// Mitsubishi GX Works2 project: 70常温静置库1130   PLC: Q10UDEH (continued)
IF NOT m_xInitial THEN
	ConveyorMotor.tLoadDelay:=T#100ms;
	ConveyorMotor.tUnloadAlarmDelay:=T#30s;
	ConveyorMotor.xPosLimit:=1;
	ConveyorMotor.xNegLimit:=1;
	ConveyorMotor.xSizeDeficientDetect:=0;
	ConveyorMotor.xZoneClear:=0;
	ConveyorMotor.tZoneClearTime:=T#10s;
	m_xInitial:=1;
END_IF;
(*//自动
//复位信号把步号置0，但xLoad与xUnload没有复位，调用程序需要注意复位后把这两个信号置零，以免发生误动作
//物料有无判断增加延时，防止开自动瞬间误动作发生*)
m_tonPresentDelay(IN:= ConveyorMotor.xCWPresent OR ConveyorMotor.xCCWPresent,
                  PT:=T#100ms,
				  Q:= m_xPresentDelay,
				  ET:= m_tPresentDelayCurrentTime);

CASE iStep OF
	0:(*//初始化*)
	ConveyorMotor.xMotorCW:=0;
	ConveyorMotor.xMotorCCW:=0;
	ConveyorMotor.iProductCategoryOut:=0;
(*	//判断物料有无传感器*)	
		IF m_xPresentDelay THEN			
			ConveyorMotor.xEmpty:=0;
			IF g_xAuto AND NOT ConveyorMotor.xError THEN(*//自动情况下进行跳转*)(*无超限报警*)
				iStep:=3;
			END_IF;
		ELSE
			ConveyorMotor.xEmpty:=1;
			IF g_xAuto AND NOT ConveyorMotor.xError THEN(*//自动情况下进行跳转*)(*无超限报警*)
				iStep:=1;	
			END_IF;		
	END_IF;	
	1: (*//上料*)
	ConveyorMotor.xNextRun:=0;
	IF ConveyorMotor.xLoad    THEN (*//上料开始*)
		ConveyorMotor.iProductCategory:=0;	(*//上料开始清除产品信息*)
		iStep:=2;		
	END_IF;
	2: (*//上料完成*)
	IF ConveyorMotor.iProductCategoryIn<>0 THEN
		ConveyorMotor.iProductCategory:=ConveyorMotor.iProductCategoryIn;(* //产品信息传入*)
	END_IF;
	IF ConveyorMotor.xloadCCW THEN
		ConveyorMotor.xMotorCCW:=1; 
		ConveyorMotor.xMotorCW:=0;
	ELSE
	    ConveyorMotor.xMotorCW:=1;  
		ConveyorMotor.xMotorCCW:=0;
	END_IF;
		m_tonLoadDelay(IN:= (ConveyorMotor.xCWPresent AND NOT ConveyorMotor.xloadCCW) 
		                                        OR (ConveyorMotor.xCCWPresent AND ConveyorMotor.xloadCCW) ,
		                               PT:= ConveyorMotor.tLoadDelay ,
		                               Q:= m_xLoadDelayOut ,
		                               ET:= m_tLoadTimer );
	    IF m_xLoadDelayOut THEN 	 
		    iStep:=3;
		END_IF;
	3:(*//下料请求*)	
	ConveyorMotor.xMotorCW:=0;
	ConveyorMotor.xMotorCCW:=0;
	ConveyorMotor.xEmpty:=0;
	IF ConveyorMotor.xUnload AND NOT ConveyorMotor.xOverWidthAlarm  THEN (*无超宽报警可以下料*)
		iStep:=4;
	END_IF;
	4:(*	//下料完成*)
	IF ConveyorMotor.xUnloadCCW THEN   
		ConveyorMotor.xMotorCCW:=1;  
		ConveyorMotor.xMotorCW:=0;
		ELSE
	    ConveyorMotor.xMotorCW:=1;  
		ConveyorMotor.xMotorCCW:=0;
	END_IF;
	ConveyorMotor.xNextRun:=1; (*下一段线体旋转*)
	ConveyorMotor.iProductCategoryOut:=ConveyorMotor.iProductCategory;(*产品型号输出给下一段线体*)
	IF NOT ConveyorMotor.xUnload THEN 
		istep:=0;
	END_IF;
END_CASE;
(*In-feed zone clear and ready to accept a load from upstream Conveyor*)
IF ldp(TRUE,g_xAuto) THEN
	m_xAutoClear:=1;
END_IF;
IF ldf(TRUE,g_xAuto) THEN
	m_xAutoClear:=0;
END_IF;
m_tonZoneClear(IN:= m_xAutoClear AND ConveyorMotor.xZoneClear ,PT:= ConveyorMotor.tZoneClearTime ,Q:=m_xZoneClearDone ,ET:= m_tZoneClearCurrentTime );
IF  m_xAutoClear AND ConveyorMotor.xZoneClear THEN
		ConveyorMotor.xMotorCW:=1; 
		iStep:=0;
END_IF;
IF ldf(TRUE, m_xAutoClear )THEN
	ConveyorMotor.xMotorCW:=0; 
END_IF;
IF NOT m_xAutoClear OR m_xZoneClearDone OR m_xPresentDelay THEN
	 m_xAutoClear:=0;
END_IF;	 
(*投入上料，搬出下料，也可用来初始化*)
IF LDP(TRUE,ConveyorMotor.xPutInto) THEN
	iStep:=0;
END_IF;
(*//当前任务显示*)
IF LDP(TRUE,ConveyorMotor.iDeviceID=g_iDeviceIDSelect) THEN
	g_iInsertTask:=ConveyorMotor.iProductCategory;
END_IF;
	(*//插入任务*)
IF g_xInsertTask AND ConveyorMotor.iDeviceID=g_iDeviceIDSelect THEN
	ConveyorMotor.iProductCategory:=g_iInsertTask;
END_IF;
(*//单线体复位，当设备号与本线体一致的时候执行复位*)
IF (g_xResetSingle AND ConveyorMotor.iDeviceID=g_iDeviceIDSelect)THEN (* //非正常情况下切断xNextRun不会复位，通过这个标志位会出发报警*)(*增加单体复位*)
	iStep:=0;
	ConveyorMotor.xNextRun:=0; 
	ConveyorMotor.xLimitAlarrm:=0;
	ConveyorMotor.xOverWidthAlarm:=0;
END_IF;
(*//手动*)
IF g_xManual THEN
(*	iStep:=0; *)(*//手动后上下料程序步骤清零*)
	(*//正转*)
	IF ConveyorMotor.xForward 
		AND ConveyorMotor.xBackward=0 
		AND ConveyorMotor.xMotorCCW=0 
		AND g_xEStop THEN
		ConveyorMotor.xMotorCW:=1;
		ConveyorMotor.xMotorCCW:=0;
		ELSE
		ConveyorMotor.xMotorCW:=0;
	END_IF;
	(*//反转*)
	IF ConveyorMotor.xBackward 
		AND ConveyorMotor.xForward=0 
		AND ConveyorMotor.xMotorCW=0 
		AND g_xEStop THEN
		ConveyorMotor.xMotorCCW:=1;
		conveyormotor.xMotorCW:=0;
		ELSE
		ConveyorMotor.xMotorCCW:=0;
	END_IF;
END_IF;
(*暂停*)
IF g_xPause THEN
	ConveyorMotor.xMotorCCW:=0;
	ConveyorMotor.xMotorCW:=0;
END_IF;
(*工作中信号输出*)
ConveyorMotor.xBusy:=ConveyorMotor.xMotorCCW OR ConveyorMotor.xMotorCW;
(*//未到达报警*)
m_tonNotArriveAlarm(IN:= iStep=0 AND ConveyorMotor.xNextRun  ,PT:= T#2s,Q:= ConveyorMotor.xNotArriveAlarm ,ET:= m_tNotArriveCurrentTime );
(*//下料超时报警*)
m_tonUnloadAlam(IN:= iStep=4,PT:=ConveyorMotor.tUnloadAlarmDelay,Q:= ConveyorMotor.xUnloadAlarm,ET:=m_tUnloadTimer );
(*//限位报警,进料检测开关失效*)
IF ( ((ConveyorMotor.xloadCCW AND NOT ConveyorMotor.xNegLimit)            (*反转上料，碰到负限位*)
	OR  ( NOT ConveyorMotor.xloadCCW AND NOT ConveyorMotor.xPosLimit)) (*正转上料，碰到正限位*)
    AND iStep=2) (*上料过程*)
    OR
   ( iStep=4 (*下料过程*)
	AND( (ConveyorMotor.xUnloadCCW AND NOT ConveyorMotor.xPosLimit)  
	OR (NOT ConveyorMotor.xUnloadCCW AND NOT ConveyorMotor.xNegLimit)))    
    THEN
    ConveyorMotor.xLimitAlarrm:=1;
    iStep:=0;
END_IF;
(*//超宽报警*)
IF (iStep=3 OR iStep=1) AND (NOT ConveyorMotor.xNegLimit OR NOT ConveyorMotor.xPosLimit) THEN
	ConveyorMotor.xOverWidthAlarm:=1;
END_IF;
(*//尺寸不足报警*)
(*//有料状态下检测两个开关都要有信号*)
IF iStep=3 AND ConveyorMotor.xSizeDeficientDetect AND (NOT ConveyorMotor.xCCWPresent OR NOT ConveyorMotor.xCWPresent)  THEN
	   ConveyorMotor.xOverWidthAlarm:=1;
	    iStep:=0;               
END_IF;
(*//总报警*)
ConveyorMotor.xError:=ConveyorMotor.xLimitAlarrm
                                              OR ConveyorMotor.xNotArriveAlarm
                                              OR ConveyorMotor.xUnloadAlarm                                             
                                              OR ConveyorMotor.xOverWidthAlarm;

(*//状态输出*)(*状态显示，容易造成指针容量不足*)
IF ConveyorMotor.xEmpty AND NOT ConveyorMotor.xBusy THEN
	m_wStateWord:=0;
END_IF;
IF ConveyorMotor.xEmpty=0 THEN
		m_wStateWord:=1;
END_IF;
IF ConveyorMotor.xBusy THEN
		m_wStateWord:=2;
END_IF;
IF ConveyorMotor.xLimitAlarrm THEN
		m_wStateWord:=3;
END_IF;
IF ConveyorMotor.xOverWidthAlarm THEN
		m_wStateWord:=4;
END_IF;
IF ConveyorMotor.xNotArriveAlarm THEN	
		m_wStateWord:=5;
END_IF;
IF ConveyorMotor.xUnloadAlarm THEN
		m_wStateWord:=6;	
END_IF;
(*选择本线体后，将状态赋值给全局变量进行显示*)
IF ConveyorMotor.iDeviceID=g_iDeviceIDSelect THEN
	g_iConveyorStatus:=m_wStateWord;
END_IF;
END_FUNCTION_BLOCK

FUNCTION_BLOCK DivideFolder
VAR_IN_OUT
  FolderIO : FolderIO;
  FolderConveyorIO : ConveyorIO;
END_VAR
VAR
  iFolderCount : INT;
  m_xInitial : BOOL;
  istep : INT;
  m_TONLoadDelay : TON;  (* 上料完成延时 *)
  m_xLoadDelay : BOOL;  (* 上料完成延时 *)
  m_tLoadDelay : TIME;  (* 上料完成延时 *)
  m_TONUpCylinderError : TON;
  m_tUpCylinderError : TIME;
  m_TONDownCylinderError : TON;
  m_tDownCylinderError : TIME;
  m_TONGrabCylinderError : TON;
  m_tGrabCylinderError : TIME;
END_VAR
VAR_INPUT
  i_xAuto : BOOL;  (* 自动 *)
END_VAR
(*拆盘机*)
(*Mr.Li修改2018.11.19调试*)
(*初始化*)
IF NOT m_xInitial  THEN
	FolderIO.i_iFloor:=3;
	 iFolderCount:=3;
	 	FolderIO.i_tSetOvertime:=T#5S;
		m_xInitial:=1;
END_IF;
(*自动*)
IF i_xAuto THEN
	FolderIO.o_xEntryPermit:=iFolderCount=3 AND FolderConveyorIO.xEmpty;(*线体状态为空且拆盘初始数量为3，才准上料*)
	m_TONLoadDelay(IN:= NOT FolderConveyorIO.xEmpty,
											PT:= T#100MS,
											Q:=m_xLoadDelay,
											ET:=m_tLoadDelay);

	CASE istep OF
		0:(*各种初始化*)
			FolderConveyorIO.xLoad:=0;
			FolderConveyorIO.xUnload:=0;
			FolderConveyorIO.xPutInto:=0;
			IF FolderConveyorIO.xEmpty THEN(*空的情况，0时上料，其他走流程*)
				IF iFolderCount=FolderIO.i_iFloor   THEN
					istep:=1; 					
				ELSE
					istep:=5;
				END_IF;	
			END_IF;		
			IF m_xLoadDelay THEN
				 IF FolderIO.i_xCylinderDownRetractDetect AND FolderIO.i_xCylinderUpRetractDetect THEN
					istep:=2;(*如果在1层，则顶起，需人为判断是否在指定位置，否则有翻框的危险*)
				ELSE
				 	istep:=3;(*如果有料不在1层，则抓紧，然后跳到第4步判断是否是叠盘，不是就放行*)
				 END_IF;
			END_IF;
		1:(*上料*)
			IF FolderIO.o_xEntryPermit THEN
				FolderConveyorIO.xLoad:=FolderIO.i_FrontConveyorNextRun;
			ELSE
				FolderConveyorIO.xLoad:=0;
			END_IF;(*有料等延时*)	
			IF m_xLoadDelay THEN
				iFolderCount:=FolderIO.i_iFloor;
				istep:=2;(**拆盘机顶起步骤*)
			END_IF;	
		2:(*上升至2层位置*)
				FolderIO.o_xCylinderDownRetract:=0;
				FolderIO.o_xCylinderDownExtend:=1;
				FolderIO.o_xCylinderUpRetract:=0;
				IF FolderIO.i_xCylinderDownExtendDetect   THEN
				istep:=3;
				END_IF;
		3:	(*夹紧夹爪*)
			IF FolderIO.i_xCylinderDownExtendDetect THEN
				FolderIO.o_xCylinderGrabExtend:=1;
				FolderIO.o_xCylinderGrabRetract:=0;
			END_IF;
			IF FolderIO.i_xCylinderGrabExtendDetect THEN
				istep:=4;
			END_IF;	
		4:(*再下降到1层，然后放行，在该位置判断是不是最后一次*)
				FolderIO.o_xCylinderUpRetract:=1;
				FolderIO.o_xCylinderUpExtend:=0;
				FolderIO.o_xCylinderDownRetract:=1;
				FolderIO.o_xCylinderDownExtend:=0;
				IF FolderIO.i_xCylinderDownRetractDetect AND FolderIO.i_xCylinderUpRetractDetect AND FolderIO.o_xExitPremit THEN
				FolderConveyorIO.xPutInto:=1;
				FolderConveyorIO.xUnload:=FolderIO.o_xExitPremit;
				ELSIF NOT FolderIO.i_xTrayDetect AND NOT FolderConveyorIO.xEmpty AND FolderIO.o_xExitPremit THEN 
						FolderConveyorIO.xUnload:=FolderIO.o_xExitPremit;
				ELSE 
					FolderConveyorIO.xPutInto:=0;
				FolderConveyorIO.xUnload:=0;
				END_IF;
					IF FolderIO.i_xCylinderDownRetractDetect AND FolderIO.i_xCylinderUpRetractDetect AND
						  FolderIO.i_xTrayDetect  AND  iFolderCount>0  AND ldp(TRUE,NOT  FolderConveyorIO.xUnload) THEN
						iFolderCount:=FolderIO.i_iFloor-1;					
					istep:=5;
					ELSIF  FolderIO.i_xCylinderDownRetractDetect AND FolderIO.i_xCylinderUpRetractDetect  AND 
						 NOT FolderIO.i_xTrayDetect   AND  FolderConveyorIO.xEmpty THEN 
						 	istep:=7;
					END_IF;

		5:(*上升到3层*)
			FolderIO.o_xCylinderUpRetract:=0;
			FolderIO.o_xCylinderUpExtend:=1;
			FolderIO.o_xCylinderDownRetract:=0;
			IF  FolderIO.i_xCylinderUpExtendDetect THEN
				istep:=6;
			END_IF;		
		6:(*松开并下降*)
			FolderIO.i_iFloor:=iFolderCount;
			IF  FolderIO.i_xCylinderUpExtendDetect  THEN
				FolderIO.o_xCylinderGrabExtend:=0;
				FolderIO.o_xCylinderGrabRetract:=1;
				IF FolderIO.i_xCylinderGrabRetractDetect THEN
					FolderIO.o_xCylinderUpRetract:=1;
					FolderIO.o_xCylinderUpExtend:=0;
					FolderIO.o_xCylinderDownRetract:=1;
					FolderIO.o_xCylinderDownExtend:=0;
				END_IF;		
			END_IF;	
			IF   FolderIO.i_xCylinderUpRetractDetect  AND FolderIO.i_xCylinderDownRetractDetect  THEN
				istep:=2;
			ELSIF iFolderCount=0 THEN 
				istep:=7;
			ELSIF  NOT FolderIO.i_xTrayDetect  THEN 
				istep:=4;
			END_IF;	
			
		7:(*恢复初始状态*)	
			FolderIO.o_xCylinderDownRetract:=1;
			FolderIO.o_xCylinderUpRetract:=1;
			FolderIO.o_xCylinderDownExtend:=0;
			FolderIO.o_xCylinderUpExtend:=0;
			FolderIO.o_xCylinderGrabExtend:=0;
			FolderIO.o_xCylinderGrabRetract:=1;
			iFolderCount:=3;
			FolderIO.i_iFloor:=3;
			IF FolderIO.i_xCylinderDownRetractDetect  AND FolderIO.i_xCylinderUpRetractDetect THEN 
			istep:=0;
			END_IF;
		END_CASE;
END_IF;(*g_xAuto那个*)	
(*手动控制气缸动作*)
		IF NOT i_xAuto THEN
			FolderIO.o_xCylinderGrabExtend:=	FolderIO.i_xCylinderGrabExtendButton;	
			FolderIO.o_xCylinderGrabRetract:=	FolderIO.i_xCylinderGrabRetractButton;	
			FolderIO.o_xCylinderUpExtend:=		FolderIO.i_xCylinderUpExtendButton;	
			FolderIO.o_xCylinderUpRetract:=		FolderIO.i_xCylinderUpRetractButton;	
			FolderIO.o_xCylinderDownExtend:=	FolderIO.i_xCylinderDownExtendButton;	
			FolderIO.o_xCylinderDownRetract:=	FolderIO.i_xCylinderDownRetractButton;		
		END_IF;
		
		(*气缸超时未到达报警，可能是没气儿漏气，也可能是开关坏了，或者气缸被卡住了*)
		m_TONGrabCylinderError(IN:= (FolderIO.o_xCylinderGrabExtend AND NOT FolderIO.i_xCylinderGrabExtendDetect) 
																OR  (FolderIO.o_xCylinderGrabRetract AND NOT FolderIO.i_xCylinderGrabRetractDetect) ,
															PT:= FolderIO.i_tSetOvertime ,Q:= FolderIO.o_xGrabCylinderError,ET:= m_tGrabCylinderError);
		m_TONDownCylinderError(IN:= (FolderIO.o_xCylinderDownExtend AND NOT FolderIO.i_xCylinderDownExtendDetect) 
																OR  (FolderIO.o_xCylinderDownRetract AND NOT FolderIO.i_xCylinderDownRetractDetect) ,
															PT:= FolderIO.i_tSetOvertime ,Q:= FolderIO.o_xDownCylinderError,ET:= m_tDownCylinderError);
		m_TONUpCylinderError(IN:= (FolderIO.o_xCylinderUpExtend AND NOT FolderIO.i_xCylinderUpExtendDetect) 
																OR  (FolderIO.o_xCylinderUpRetract AND NOT FolderIO.i_xCylinderUpRetractDetect) ,
															PT:= FolderIO.i_tSetOvertime ,Q:= FolderIO.o_xUpCylinderError,ET:= m_tUpCylinderError);
		
		
(*手动恢复程序，不要自动恢复，因为自动恢复需要检测传感器，有可能引起误动作*)		
IF NOT  i_xAuto
	THEN istep:=FolderIO.m_iStepInput;
				iFolderCount:=FolderIO.m_CountInput;
END_IF;(*使用拆盘机时，当拆盘小于3盘时恢复尽量从第2步开始恢复，既先手动松开夹爪，将货物降到第1层，然后将步骤跳到第2步，在将数量填入当前拆盘机剩余的盘数，然后切换成自动即可*)
END_FUNCTION_BLOCK

FUNCTION_BLOCK FanucRobot
VAR_IN_OUT
  FanucRobotIO : FanucRobotIO;
END_VAR
VAR
  m_iSNO : INT;
  m_xPNSPass : BOOL;  (* 收到程序号 *)
  m_tonStartDelay : TON;  (* 启动延时 *)
  m_xStartDelay : BOOL;
  m_tStartDelayCurrentTime : TIME;
END_VAR
(***********************************************************
发那科机器人自动启动程序


***********************************************************)

(*无自动状态，示教盒处于本地状态，把各标志位复位*)
IF FanucRobotIO.i_xTPENBL AND NOT g_xAuto THEN
	FanucRobotIO.o_xPNSTROBE:=0;
	FanucRobotIO.o_xCSTOPI:=0;
	FanucRobotIO.o_xPROD_START:=0;
	FanucRobotIO.o_xRESET:=0;
END_IF;
(*远程模式*)
IF g_xAuto THEN
	FanucRobotIO.o_xREMOTE:=1;
	ELSE
	FanucRobotIO.o_xREMOTE:=0;
END_IF;
(*程序启动后复位启动标志位*)
IF FanucRobotIO.i_xPROG_RUN AND FanucRobotIO.i_xBUSY THEN
	FanucRobotIO.i_xCommandStart:=0;
END_IF;
(*示教盒旋清除报警*)
IF ldf(TRUE,FanucRobotIO.i_xTPENBL)THEN
	FanucRobotIO.o_xRESET:=1;
	FanucRobotIO.o_xCSTOPI:=1;
END_IF;
(*启动程序号条件*)
IF FanucRobotIO.i_xSYSRDY 
	AND FanucRobotIO.i_xCMDENBL
	AND FanucRobotIO.i_xCommandStart
	AND NOT FanucRobotIO.i_xPROG_RUN 
	AND NOT FanucRobotIO.i_xBUSY THEN
	FanucRobotIO.o_xRESET:=0;
	FanucRobotIO.o_xCSTOPI:=0;
	IF FanucRobotIO.i_iMotionNumber <> 0 (*只要动作编号不为0，就给他信号*)
		AND NOT FanucRobotIO.o_xPNSTROBE THEN
		FanucRobotIO.o_xPNSTROBE:=1;
		FanucRobotIO.o_xPROD_START:=1;
		FanucRobotIO.o_iPNS:=FanucRobotIO.i_iMotionNumber;(*并把任务号传给他*)
	END_IF;
	(*程序号校验*)
	IF FanucRobotIO.i_xSNACK THEN(*数据传回之后再校验*)
		m_iSNO:=BITARR_TO_INT(FanucRobotIO.i_arrxSNO[0] , 8 );
		IF m_iSNO=FanucRobotIO.o_iPNS THEN
			m_xPNSPass:=1;(*校验成功,等100MS复位Start信号*)
			FanucRobotIO.o_xPNSTROBE:=0;
		ELSE
			FanucRobotIO.o_xPNSFailed:=1;(*校验失败*)
			FanucRobotIO.o_xPROD_START:=0;(*立刻复位，不生成任务*)
		END_IF;
	END_IF;
END_IF;
m_tonStartDelay(IN:= m_xPNSPass ,PT:= T#100ms ,Q:= m_xStartDelay ,ET:=m_tStartDelayCurrentTime );
IF m_xStartDelay THEN
	FanucRobotIO.o_xPROD_START:=0;
	FanucRobotIO.i_xCommandStart:=0;
	m_xPNSPass:=0;
END_IF;
END_FUNCTION_BLOCK

FUNCTION_BLOCK Folder
VAR_IN_OUT
  FolderIO : FolderIO;
END_VAR
VAR
  m_xInitial : BOOL;
END_VAR
VAR_IN_OUT
  FolderConveyorIO : ConveyorIO;
END_VAR
VAR
  iFolderCount : INT;
  istep : INT;
  m_TONLoadDelay : TON;  (* 上料完成延时 *)
  m_xLoadDelay : BOOL;  (* 上料完成延时 *)
  m_tLoadDelay : TIME;  (* 上料完成延时 *)
  m_TONUpCylinderError : TON;
  m_tUpCylinderError : TIME;
  m_TONDownCylinderError : TON;
  m_tDownCylinderError : TIME;
  m_TONGrabCylinderError : TON;
  m_tGrabCylinderError : TIME;
END_VAR
VAR_INPUT
  i_xAuto : BOOL;  (* 自动 *)
  i_xManual : BOOL;  (* 手动 *)
END_VAR
(*叠盘机*)
(*sb刘写的*)
(*初始化*)
(*18/11/17 YAOBO更改*)
(*增加允许下料信号o_xExitPrimit，码垛完成后给允许下料第7步给出*)
(*18/11/28 YAOBO更改*)
(*增加叠盘个数输出FolderIO.o_CountResponsPC*)
IF NOT m_xInitial THEN
	FolderIO.i_iFloor:=3;
	FolderIO.i_tSetOvertime:=T#5S;
	
	m_xInitial:=1;
END_IF;
(*自动*)
FolderIO.o_xEntryPermit:=FolderConveyorIO.xEmpty;(*叠盘机的话，只要空了，就允许上料，拆盘则是拆完才允许*)
IF i_xAuto THEN
				m_TONLoadDelay(IN:= NOT FolderConveyorIO.xEmpty,
													PT:= T#100MS,
													Q:=m_xLoadDelay,
													ET:=m_tLoadDelay);
	CASE istep OF
		0:(*各种初始化*)
			FolderConveyorIO.xLoad:=0;
			FolderConveyorIO.xUnload:=0;
			FolderConveyorIO.xPutInto:=0;
			FolderIo.o_xExitPremit:=0;	
			IF (*0 AND*)  FolderConveyorIO.xEmpty THEN
				istep:=1;(*空着就去1上料*)
			END_IF;	
			IF 0 AND    m_xLoadDelay  THEN(*if 有料*)
				IF  FolderIO.i_xCylinderDownExtendDetect  AND FolderIO.i_xCylinderUpExtendDetect  THEN(*if 在下层*)
					IF iFolderCount=FolderIO.i_iFloor THEN(*if 是最后一次*)
						istep:=7;
					ELSE(*不是最后一次去5，是就去7*)
						istep:=5;
					END_IF;(*if 是最后一次*)	
				ELSE(*不在下层去2*)
				istep:=2;
				END_IF;	(*if 在下层*)			
			END_IF;(*if 有料*)
			
		1:(*上料*)
			IF FolderIO.i_xEntryEnable THEN
				FolderConveyorIO.xLoad:=1;
			ELSE
				FolderConveyorIO.xLoad:=0;
			END_IF;(*not Empty了等个延时*)	

			IF (*0 AND*)   m_xLoadDelay  AND (iFolderCount>0 AND iFolderCount<FolderIO.i_iFloor) AND FolderIO.i_xFolderEnable THEN
				istep:=2;
			ELSIF (*0 AND*)   m_xLoadDelay AND iFolderCount=0 AND FolderIO.i_xFolderEnable THEN(*=0表示是第一次，第一次直接抓紧上升*)
				istep:=5;	
			END_IF;	
		2:(*下降，到2层位置*)
				FolderIO.o_xCylinderUpRetract:=0;
				FolderIO.o_xCylinderUpExtend:=1;
				FolderIO.o_xCylinderDownRetract:=1;
				FolderIO.o_xCylinderDownExtend:=0;
				IF FolderIO.i_xCylinderUpExtendDetect AND NOT FolderIO.i_xCylinderDownExtendDetect THEN
					istep:=3;
				END_IF;
		3:	(*松开夹爪*)
			IF FolderConveyorIO.xCWPresent AND NOT FolderConveyorIO.xEmpty THEN(*有感应到才松开*)
				FolderIO.o_xCylinderGrabExtend:=0;
				FolderIO.o_xCylinderGrabRetract:=1;
				IF (*0 AND*)   FolderIO.i_xCylinderGrabRetractDetect THEN
					IF iFolderCount=FolderIO.i_iFloor-1 THEN
						iFolderCount:=FolderIO.i_iFloor;(*最后一次到这里就刷新计数，方便故障恢复*)
					END_IF;	
					istep:=4;
				END_IF;	
			END_IF;	
		4:(*再下降，去1层*)
				FolderIO.o_xCylinderUpRetract:=0;
				FolderIO.o_xCylinderUpExtend:=1;
				FolderIO.o_xCylinderDownRetract:=0;
				FolderIO.o_xCylinderDownExtend:=1;
				IF FolderIO.i_xCylinderDownExtendDetect  AND FolderIO.i_xCylinderUpExtendDetect  THEN
					IF iFolderCount<FolderIO.i_iFloor-1 THEN
						istep:=5;
					ELSE
						istep:=7;
					END_IF;	
				END_IF;		
		5:(*抓紧*)
			IF FolderIO.i_xCylinderDownExtendDetect  AND FolderIO.i_xCylinderUpExtendDetect  THEN
				FolderIO.o_xCylinderGrabExtend:=1;
				FolderIO.o_xCylinderGrabRetract:=0;
				IF (*0 AND*)   FolderIO.i_xCylinderGrabExtendDetect THEN
					iFolderCount:=iFolderCount+1;
					istep:=6;
				END_IF;	
			END_IF;		
		6:(*上升到3层*)
			FolderIO.o_xCylinderUpRetract:=1;
			FolderIO.o_xCylinderUpExtend:=0;
			FolderIO.o_xCylinderDownRetract:=1;
			FolderIO.o_xCylinderDownExtend:=0;
			IF (*0 AND *)  FolderIO.i_xCylinderDownRetractDetect AND FolderIO.i_xCylinderUpRetractDetect THEN
				FolderConveyorIO.xPutInto:=1;(*刷新成Empty的*)
				istep:=0;
			END_IF;
		7:(*下料*)
		FolderIo.o_xExitPremit:=1;	(*给出允许下料信号*)
		FolderConveyorIO.xUnload:=	FolderIO.i_xExitEnable AND FolderIO.i_xCylinderGrabRetractDetect;(*给下料信号，不要刷新完成*)
	(*			IF	FolderIO.i_xExitEnable AND FolderIO.i_xCylinderGrabRetractDetect	THEN(*保证不会挂到叉手*)
(*				FolderConveyorIO.xUnload:=1;
			ELSE
				FolderConveyorIO.xPutInto:=1;(*刷新成Empty的*)
	(*			FolderConveyorIO.xUnload:=0;
			END_IF;	*)
			IF FolderConveyorIO.xEmpty THEN(*确保空了才回0，不然还在这里等Unload信号*)
				iFolderCount:=0;
				istep:=0;
			END_IF;	 
		END_CASE;
END_IF;(*g_xAuto那个*)	
(*手动控制气缸动作*)
		IF i_xManual THEN
			FolderIO.o_xCylinderGrabExtend:=	FolderIO.i_xCylinderGrabExtendButton;	
			FolderIO.o_xCylinderGrabRetract:=	FolderIO.i_xCylinderGrabRetractButton;	
			FolderIO.o_xCylinderUpExtend:=		FolderIO.i_xCylinderUpExtendButton;	
			FolderIO.o_xCylinderUpRetract:=		FolderIO.i_xCylinderUpRetractButton;	
			FolderIO.o_xCylinderDownExtend:=	FolderIO.i_xCylinderDownExtendButton;	
			FolderIO.o_xCylinderDownRetract:=	FolderIO.i_xCylinderDownRetractButton;		
		END_IF;
		
		(*气缸超时未到达报警，可能是没气儿漏气，也可能是开关坏了，或者气缸被卡住了*)
		m_TONGrabCylinderError(IN:= (FolderIO.o_xCylinderGrabExtend AND NOT FolderIO.i_xCylinderGrabExtendDetect) 
																OR  (FolderIO.o_xCylinderGrabRetract AND NOT FolderIO.i_xCylinderGrabRetractDetect) ,
															PT:= FolderIO.i_tSetOvertime ,Q:= FolderIO.o_xGrabCylinderError,ET:= m_tGrabCylinderError);
		m_TONDownCylinderError(IN:= (FolderIO.o_xCylinderDownExtend AND NOT FolderIO.i_xCylinderDownExtendDetect) 
																OR  (FolderIO.o_xCylinderDownRetract AND NOT FolderIO.i_xCylinderDownRetractDetect) ,
															PT:= FolderIO.i_tSetOvertime ,Q:= FolderIO.o_xDownCylinderError,ET:= m_tDownCylinderError);
		m_TONUpCylinderError(IN:= (FolderIO.o_xCylinderUpExtend AND NOT FolderIO.i_xCylinderUpExtendDetect) 
																OR  (FolderIO.o_xCylinderUpRetract AND NOT FolderIO.i_xCylinderUpRetractDetect) ,
															PT:= FolderIO.i_tSetOvertime ,Q:= FolderIO.o_xUpCylinderError,ET:= m_tUpCylinderError);
		
	FolderIO.o_CountResponsPC:= iFolderCount;(*叠盘数量输出*)
IF NOT  i_xAuto
	THEN istep:=FolderIO.m_iStepInput;
				iFolderCount:=FolderIO.m_CountInput;
END_IF;(*使用第1种叠盘机时，当叠盘小于3盘时，恢复尽量从第4步开始恢复，既先手动松开夹爪，将货物降到第1层，然后将步骤跳到第4步，在将数量填入当前叠盘机所叠的盘数-1，然后切换成自动即可
					若是实际叠盘数量为3，则步骤 跳到7，数量填3*)
END_FUNCTION_BLOCK

FUNCTION_BLOCK FolderII
VAR_IN_OUT
  FolderIO : FolderIO;
  FolderConveyorIO : ConveyorIO;
END_VAR
VAR_INPUT
  i_xAuto : BOOL;  (* 自动 *)
END_VAR
VAR
  iFolderCount : INT;
  m_xInitial : BOOL;
  istep : INT;
  m_TONLoadDelay : TON;  (* 上料完成延时 *)
  m_xLoadDelay : BOOL;  (* 上料完成延时 *)
  m_tLoadDelay : TIME;  (* 上料完成延时 *)
  m_TONUpCylinderError : TON;
  m_tUpCylinderError : TIME;
  m_TONDownCylinderError : TON;
  m_tDownCylinderError : TIME;
  m_TONGrabCylinderError : TON;
  m_tGrabCylinderError : TIME;
END_VAR
VAR_INPUT
  i_xManual : BOOL;  (* 手动 *)
END_VAR
(*叠盘机II型*)
(*初始化*)
(*18/11/17 YAOBO更改*)
(*增加允许下料信号o_xExitPrimit，码垛完成后给允许下料第7步给出*)
IF NOT m_xInitial THEN
	FolderIO.i_iFloor:=3;
	FolderIO.i_tSetOvertime:=T#5S;
	
	m_xInitial:=1;
END_IF;
(*自动*)
FolderIO.o_xEntryPermit:=FolderConveyorIO.xEmpty;(*叠盘机的话，只要空了，就允许上料，拆盘则是拆完才允许*)
IF i_xAuto THEN
				m_TONLoadDelay(IN:= NOT FolderConveyorIO.xEmpty,
													PT:= T#100MS,
													Q:=m_xLoadDelay,
													ET:=m_tLoadDelay);
	CASE istep OF
		0:(*各种初始化*)
			FolderConveyorIO.xLoad:=0;
			FolderConveyorIO.xUnload:=0;
			FolderConveyorIO.xPutInto:=0;
			FolderIo.o_xExitPremit:=0;	
			FolderIo.i_xExitEnable:=0;
			IF (*0 AND*)  FolderConveyorIO.xEmpty THEN
				istep:=1;(*空着就去1上料*)
			END_IF;	
			IF 0 AND    m_xLoadDelay  THEN(*if 有料*)
				IF  FolderIO.i_xCylinderDownRetractDetect  AND FolderIO.i_xCylinderUpRetractDetect  THEN(*if 在下层*)
					IF iFolderCount=FolderIO.i_iFloor THEN(*if 是最后一次*)
						istep:=7;
					ELSE(*不是最后一次去5，是就去7*)
						istep:=5;
					END_IF;(*if 是最后一次*)	
				ELSE(*不在下层去2*)
				istep:=2;
				END_IF;	(*if 在下层*)			
			END_IF;(*if 有料*)
			
		1:(*上料*)
			IF FolderIO.i_xEntryEnable THEN
				FolderConveyorIO.xLoad:=1;
			ELSE
				FolderConveyorIO.xLoad:=0;
			END_IF;(*not Empty了等个延时*)	

			IF (*0 AND*)   m_xLoadDelay  AND (iFolderCount>0 AND iFolderCount<FolderIO.i_iFloor) AND FolderIO.i_xFolderEnable THEN
				istep:=2;
			ELSIF (*0 AND*)   m_xLoadDelay AND iFolderCount=0 AND FolderIO.i_xFolderEnable THEN(*=0表示是第一次，第一次直接抓紧上升*)
				istep:=4;	
			END_IF;	
		2:(*上升，到2层位置*)
				FolderIO.o_xCylinderUpRetract:=0;
				FolderIO.o_xCylinderUpExtend:=0;
				FolderIO.o_xCylinderDownRetract:=0;
				FolderIO.o_xCylinderDownExtend:=1;
				IF   FolderIO.i_xCylinderDownExtendDetect THEN
					istep:=3;
				END_IF;
		3:	(*松开夹爪,并降到1层*)
			IF  FolderIO.i_xTrayDetect AND NOT FolderConveyorIO.xEmpty THEN(*有感应到才松开*)
				FolderIO.o_xCylinderGrabExtend:=0;
				FolderIO.o_xCylinderGrabRetract:=1;
				IF (*0 AND*)   FolderIO.i_xCylinderGrabRetractDetect THEN
					FolderIO.o_xCylinderDownRetract:=1;
					FolderIO.o_xCylinderDownExtend:=0;
					IF iFolderCount=FolderIO.i_iFloor-1 THEN
						iFolderCount:=FolderIO.i_iFloor;(*最后一次到这里就刷新计数，方便故障恢复*)
					END_IF;	
					IF FolderIO.i_xCylinderDownRetractDetect  THEN 
					istep:=4;
					END_IF;
				END_IF;	
			END_IF;	
		4:(*再上升，去3层*)
		IF iFolderCount<FolderIO.i_iFloor-1 THEN 
				FolderIO.o_xCylinderUpRetract:=0;
				FolderIO.o_xCylinderUpExtend:=1;
				FolderIO.o_xCylinderDownRetract:=0;
				FolderIO.o_xCylinderDownExtend:=0;
				IF  FolderIO.i_xCylinderUpExtendDetect
					THEN  istep:=5;
				END_IF;
		ELSE FolderIO.o_xCylinderUpRetract:=1;
				FolderIO.o_xCylinderUpExtend:=0;
				FolderIO.o_xCylinderDownRetract:=1;
				FolderIO.o_xCylinderDownExtend:=0;
				   IF  FolderIO.i_xCylinderUpRetractDetect AND FolderIO.i_xCylinderDownRetractDetect THEN 
				   	 istep:=7;
				   END_IF;
		END_IF;
			
	
		5:(*抓紧*)
			IF  FolderIO.i_xCylinderUpExtendDetect  THEN
				FolderIO.o_xCylinderGrabExtend:=1;
				FolderIO.o_xCylinderGrabRetract:=0;
				IF (*0 AND*)   FolderIO.i_xCylinderGrabExtendDetect THEN
					iFolderCount:=iFolderCount+1;
					istep:=6;
				END_IF;	
			END_IF;		
		6:(*下降到1层*)
			FolderIO.o_xCylinderUpRetract:=1;
			FolderIO.o_xCylinderUpExtend:=0;
			FolderIO.o_xCylinderDownRetract:=1;
			FolderIO.o_xCylinderDownExtend:=0;
			IF (*0 AND *)  FolderIO.i_xCylinderDownRetractDetect AND FolderIO.i_xCylinderUpRetractDetect THEN
				FolderConveyorIO.xPutInto:=1;(*刷新成Empty的*)
				istep:=0;
			END_IF;
		7:(*下料*)
		FolderIo.o_xExitPremit:=1;	(*给出允许下料信号*)
		IF FolderIo.o_xExitPremit
			THEN FolderIo.i_xExitEnable:=1;
		END_IF;
		FolderConveyorIO.xUnload:=	FolderIO.i_NextConveyorEmpty AND FolderIO.i_xCylinderGrabRetractDetect AND
		 FolderIO.i_xCylinderDownRetractDetect AND FolderIO.i_xCylinderUpRetractDetect ;(*给下料信号，不要刷新完成*)
	(*			IF	FolderIO.i_xExitEnable AND FolderIO.i_xCylinderGrabRetractDetect	THEN(*保证不会挂到叉手*)
(*				FolderConveyorIO.xUnload:=1;
			ELSE
				FolderConveyorIO.xPutInto:=1;(*刷新成Empty的*)
	(*			FolderConveyorIO.xUnload:=0;
			END_IF;	*)
			IF FolderConveyorIO.xEmpty THEN(*确保空了才回0，不然还在这里等Unload信号*)
				iFolderCount:=0;
				istep:=0;
			END_IF;	 
		END_CASE;
END_IF;(*g_xAuto那个*)	
(*手动控制气缸动作*)
		IF i_xManual THEN
			FolderIO.o_xCylinderGrabExtend:=	FolderIO.i_xCylinderGrabExtendButton;	
			FolderIO.o_xCylinderGrabRetract:=	FolderIO.i_xCylinderGrabRetractButton;	
			FolderIO.o_xCylinderUpExtend:=		FolderIO.i_xCylinderUpExtendButton;	
			FolderIO.o_xCylinderUpRetract:=		FolderIO.i_xCylinderUpRetractButton;	
			FolderIO.o_xCylinderDownExtend:=	FolderIO.i_xCylinderDownExtendButton;	
			FolderIO.o_xCylinderDownRetract:=	FolderIO.i_xCylinderDownRetractButton;		
		END_IF;
		
		(*气缸超时未到达报警，可能是没气儿漏气，也可能是开关坏了，或者气缸被卡住了*)
		m_TONGrabCylinderError(IN:= (FolderIO.o_xCylinderGrabExtend AND NOT FolderIO.i_xCylinderGrabExtendDetect) 
																OR  (FolderIO.o_xCylinderGrabRetract AND NOT FolderIO.i_xCylinderGrabRetractDetect) ,
															PT:= FolderIO.i_tSetOvertime ,Q:= FolderIO.o_xGrabCylinderError,ET:= m_tGrabCylinderError);
		m_TONDownCylinderError(IN:= (FolderIO.o_xCylinderDownExtend AND NOT FolderIO.i_xCylinderDownExtendDetect) 
																OR  (FolderIO.o_xCylinderDownRetract AND NOT FolderIO.i_xCylinderDownRetractDetect) ,
															PT:= FolderIO.i_tSetOvertime ,Q:= FolderIO.o_xDownCylinderError,ET:= m_tDownCylinderError);
		m_TONUpCylinderError(IN:= (FolderIO.o_xCylinderUpExtend AND NOT FolderIO.i_xCylinderUpExtendDetect) 
																OR  (FolderIO.o_xCylinderUpRetract AND NOT FolderIO.i_xCylinderUpRetractDetect) ,
															PT:= FolderIO.i_tSetOvertime ,Q:= FolderIO.o_xUpCylinderError,ET:= m_tUpCylinderError);
		
(*手动恢复程序，不要自动恢复，因为自动恢复需要检测传感器，有可能引起误动作*)		
IF NOT  i_xAuto
	THEN istep:=FolderIO.m_iStepInput;
				iFolderCount:=FolderIO.m_CountInput;
END_IF;(*使用第2种叠盘机时，当叠盘小于3盘时，恢复尽量从第4步开始恢复，既先手动松开夹爪，将货物降到第1层，然后将步骤跳到第4步，在将数量填入当前叠盘机所叠的盘数-1，然后切换成自动即可
					若是实际叠盘数量为3，则步骤 跳到7，数量填3*)
(*给上位机叠盘数量*)
IF istep=1 AND  iFolderCount=0 THEN 
		FolderIO.o_CountResponsPC:=0;
ELSIF  istep=6 AND   iFolderCount=1 THEN 
		FolderIO.o_CountResponsPC:=1;
ELSIF  istep=6 AND   iFolderCount=2 THEN 
		FolderIO.o_CountResponsPC:=2;
ELSIF  istep=3 AND   iFolderCount=2 THEN 
		 FolderIO.o_CountResponsPC:=3;
END_IF;

IF FolderIO.i_FrontConveyorTypeInfo=2 OR istep=7(*不同批次或者叠满后给上位机出料请求*)
		THEN FolderIO.o_RequestPC:=2;
END_IF;
IF FolderIO.i_FrontConveyorTypeInfo=2 THEN(*当不同批次时，步骤跳到7*)
		 istep:=7;
END_IF;
END_FUNCTION_BLOCK

FUNCTION_BLOCK PackCommunication
VAR_IN_OUT
  ConveyorIO : ConveyorIO;
  PackCommunicationIO : PackCommunicationIO;
  FanucRobotIO : FanucRobotIO;
END_VAR
VAR_OUTPUT
  o_iErrorNub : INT;
  o_xReqSuccess : BOOL;
END_VAR
VAR
  m_xReqSuccess : BOOL;
  m_iStep : INT;
  m_arrwCode : ARRAY [1..8] OF BatteryCode;
END_VAR
VAR_INPUT
  i_arrxPresentDetect : ARRAY [1..8] OF BOOL;
END_VAR
VAR
  m_iCoordinateX : INT;
  m_iCoordinateY : INT;
  m_arriPresentDetect : ARRAY [1..8] OF INT;
  ii : INT;
END_VAR
VAR CONSTANT
  MAX_ROW : INT := 8;
  MAX_COLUMN : INT := 8;
END_VAR
VAR
  m_xSupplement : BOOL;
END_VAR
VAR CONSTANT
  ROW_TIMES : INT := 1;
  GET_QUANTITY : INT := 8;
END_VAR
VAR
  m_iRowReminder : INT;
  m_xEno : BOOL;
  m_iRowReminderTemp : INT;
END_VAR
(***************************************************************************)
(*
DB1区(PC->PLC)10个字		
"字(16位）序号
(从1开始)"	功能描述	具体参数解释
1	请求确认	"1：复位
2：读码(入库申请）成功
101：条码空
102：条码规则校验失败
103：步号校验失败
"
2	放行	"1：复位
2：完成,放行
3：撤销完成 "
3	单次装载应答	"1：复位
2：允许开始"
4	单次装载处理完成	"1：复位
2：完成
3：电芯为空"
)*
DB2区(PLC->PC)200个字		
"字(16位）序号
(从1开始)"	功能描述	具体参数解释
1	装载请求	"１：复位
２：请求"
2	装载全部完成	"1：复位
2：请求 "
3	单次装载请求	"1：复位
2：请求 "
4	单次装载完成	"1：复位
2：完成"
5	行坐标	从1开始
6	列坐标	从1开始
7	电芯码(15*11=165)	"电芯码24字符，
占12个字，加上预留的每个分配15个字"

顺序执行步骤
0  初始化
1  框码扫码请求
2  单次抓取请求
3  整排抓取
4  补料
5  完成


(***************************************************************************)
m_iRowReminder:= ( m_iCoordinateX-1 MOD GET_QUANTITY )+1;(*//通过位置与抓取数量取余数，判断是否的抓取位置为一排的最后一个*)
CASE m_iStep OF
	0:;(*//初始化*)
	m_iStep:=1;
	1:(*发送框码的扫码请求*)
	IF NOT ConveyorIO.xEmpty AND NOT FanucRobotIO.io_xMutexLock THEN
		PackCommunicationIO.o_iRequestPLCPC:=2;
		ELSE
		PackCommunicationIO.o_iRequestPLCPC:=1;
	END_IF;
	(*//请求确认*)
	CASE PackCommunicationIO.i_iResponsPCPLC OF 
		0:;
		1:;(*//复位*)
		2:(*//读码（入库申请）成功*)
		m_iStep:=2;
		m_xSupplement:=0;
		m_iCoordinateX:=1;(*//框码扫码成功后把坐标改为1,1*)
		m_iCoordinateY:=1;
		FanucRobotIO.io_xMutexLock:=1;
		3:(*//取放货完成*)
		ConveyorIO.xPutInto:=1; 
		4:(*//旋转*)
		;
		5:(*//不旋转*)
		;
		101:(*//条码空*)
		o_iErrorNub:=101;
		m_iStep:=0;
		102:(*//条码规则检验失败*)
		o_iErrorNub:=102;
		m_iStep:=0;
		103:(*//步号校验失败*)
		o_iErrorNub:=103;
		m_iStep:=0;
		104:(*//无库位可用*)
		o_iErrorNub:=104;
		m_iStep:=0;
	END_CASE;
	2:(*//单次抓取请求，分为单次多个产品抓取与补料程序*)
	IF FanucRobotIO.i_xSYSRDY 
		AND NOT FanucRobotIO.i_xBUSY
		AND NOT FanucRobotIO.i_xPROG_RUN
		AND i_arrxPresentDetect[1] 
		AND PackCommunicationIO.i_iSinglePackResponsePCPLC=1 THEN(*//机器人准备就绪、组装下线有料*)
		PackCommunicationIO.o_iSinglePackRequestPLCPC:=2;
	END_IF;
	IF (*LDP(TRUE,PackCommunicationIO.i_iSinglePackResponsePCPLC=2)*) PackCommunicationIO.i_iSinglePackResponsePCPLC=2 THEN(*//请求成功*)
		PackCommunicationIO.o_iSinglePackRequestPLCPC:=1;(*//复位请求*)
		IF m_xSupplement THEN(*//补料标志位，为1进行补料操作，为0进行整排抓取*)
			m_iStep:=4;(*//补料*)
			ELSE
		 	m_iStep:=3;(*//整排抓取*)
			FOR ii:=1 TO GET_QUANTITY BY 1 DO(*//记录哪个位置缺料*)
				IF i_arrxPresentDetect[ii] THEN(*//传感器检测*)
 m_arriPresentDetect[ii]:=0;
 ELSE
 m_arriPresentDetect[ii]:=ii;(*//记录缺料的位置*)
				END_IF;
			END_FOR;
		END_IF;
	END_IF;
	3:  (*//整排抓取*)
	FanucRobotIO.o_iPNS:=10101;(*//步骤号*)
	FanucRobotIO.o_uiOffset_X:=m_iCoordinateX;
	FanucRobotIO.o_uiOffset_Y:=m_iCoordinateY;
	PackCommunicationIO.o_iXCoordinatePLCPC:=m_iCoordinateX;(*//放置位置发送给上位机*)
	PackCommunicationIO.o_iYCoordinatePLCPC:=m_iCoordinateY;	
	IF LDF(TRUE,FanucRobotIO.i_xBUSY OR FanucRobotIO.i_xPROG_RUN) THEN(*//抓取动作完成*)
		FOR ii:=1 TO GET_QUANTITY BY 1 DO (*//判断有无补料信息*)
			IF m_arriPresentDetect[ii]<>0  THEN(*//有补料*)(*//补料不是最后一个的算法*)
				m_iCoordinateX:=m_arriPresentDetect[ii]+((m_iCoordinateX-1)/GET_QUANTITY)*GET_QUANTITY;
				m_xSupplement:=1;
				m_iStep:=2;(*//有补料*)
				EXIT;
			END_IF;			
		END_FOR;
		IF ii=GET_QUANTITY+1  THEN  (*//无补料*)
			m_xSupplement:=0;
			IF m_iCoordinateY = MAX_ROW (*//达到最大列*)
				AND ((m_iCoordinateX-1)/GET_QUANTITY+1=ROW_TIMES) 
				THEN(*//偏移量为最大的值时,排抓取为最后一排*)
				m_iStep:=5;(*//装盘完成*)
				ELSE
				m_iStep:=2;(*//请求下一次装盘*)			
				IF (m_iCoordinateX-1)/GET_QUANTITY+1=ROW_TIMES THEN
 m_iCoordinateX:=1;                                              (*//开始执行下一列*)
 m_iCoordinateY:=m_iCoordinateY+1;
 ELSE
 m_iCoordinateX:=((m_iCoordinateX-1)/GET_QUANTITY+1)*GET_QUANTITY+1;
				END_IF;
			END_IF;
		END_IF;
	END_IF;
	4: (*//补料*)
	FanucRobotIO.o_iPNS:=10102;(*//步骤号*)
	FanucRobotIO.o_uiOffset_X:=m_iCoordinateX;
	FanucRobotIO.o_uiOffset_Y:=m_iCoordinateY;
	PackCommunicationIO.o_iXCoordinatePLCPC:=m_iCoordinateX;(*//放置位置发送给上位机*)
	PackCommunicationIO.o_iYCoordinatePLCPC:=m_iCoordinateY;
	IF LDF(TRUE,FanucRobotIO.i_xBUSY OR FanucRobotIO.i_xPROG_RUN) THEN(*//抓取动作完成*)
		FOR ii:=m_iRowReminder+1 TO GET_QUANTITY BY 1 DO (*//判断有无补料信息*)
			IF m_arriPresentDetect[ii]<>0  THEN(*//有补料*)(*//补料不是最后一个的算法*)
				m_iCoordinateX:=m_arriPresentDetect[ii]+((m_iCoordinateX-1)/GET_QUANTITY)*GET_QUANTITY;
				m_xSupplement:=1;
				m_iStep:=2;(*//有补料*)
				EXIT;
			END_IF;	
		END_FOR;
		IF ii=GET_QUANTITY+1  THEN  (*//无补料*)
			m_xSupplement:=0;
			IF m_iCoordinateY = MAX_ROW (*//达到最大列*)
				AND ((m_iCoordinateX-1)/GET_QUANTITY+1=ROW_TIMES)
				THEN(*//偏移量为最大的值时,排抓取为最后一排*)
				m_iStep:=5;(*//装盘完成*)
				ELSE
				m_iStep:=2;(*//请求下一次装盘*)			
				IF (m_iCoordinateX-1)/GET_QUANTITY+1=ROW_TIMES THEN
 m_iCoordinateX:=1;                                              (*//开始执行下一列*)
 m_iCoordinateY:=m_iCoordinateY+1;
 ELSE
 m_iCoordinateX:=((m_iCoordinateX-1)/GET_QUANTITY+1)*GET_QUANTITY+1;(*//这一列继续往后排*)
				END_IF;
			END_IF;
		END_IF;
	END_IF;
	5: (*//完成*)
	PackCommunicationIO.o_iSinglePackDonePLCPC:=2;
	IF PackCommunicationIO.i_iSinglePackDoneAknPCPLC =2 THEN
		PackCommunicationIO.o_iSinglePackDonePLCPC:=1;
		m_iCoordinateX:=1;